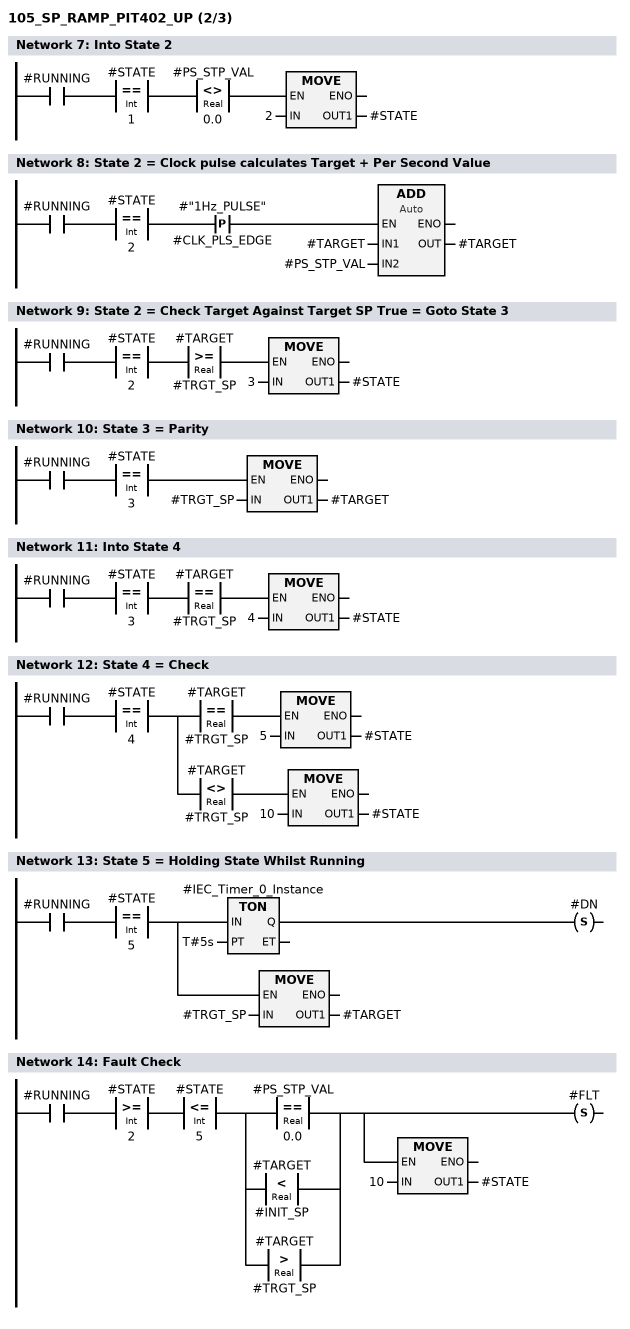
   RUNG wire#powerrail
      Contact( #RUNNING )
      { S7_Templates := "SrcType := Int" } EQ_Contact(in1 := #STATE, in2 := 1)
      { S7_Templates := "SrcType := Real" } NE_Contact(in1 := #PS_STP_VAL, in2 := 0.0)
      Move(in := 2, out1 => #STATE)
   END_RUNG
   // the same network as SCL:
   IF #RUNNING AND (#STATE = 1) AND (#PS_STP_VAL <> 0.0) THEN #STATE := 2; END_IF;
END_REGION

REGION Network 8: State 2 = Clock pulse calculates Target + Per Second Value
   RUNG wire#powerrail
      Contact( #RUNNING )
      { S7_Templates := "SrcType := Int" } EQ_Contact(in1 := #STATE, in2 := 2)
      P_Contact(operand := #"1Hz_PULSE", bit := #CLK_PLS_EDGE)
      Add(in1 := #TARGET, in2 := #PS_STP_VAL, out => #TARGET)
   END_RUNG
   // the same network as SCL:
   #_w1 := #RUNNING AND (#STATE = 2) AND #"1Hz_PULSE" AND NOT #CLK_PLS_EDGE;   // rising edge of #"1Hz_PULSE"
   #CLK_PLS_EDGE := #"1Hz_PULSE";
   IF #_w1 THEN #TARGET := #TARGET + #PS_STP_VAL; END_IF;
END_REGION

REGION Network 9: State 2 = Check Target Against Target SP True = Goto State 3
   RUNG wire#powerrail
      Contact( #RUNNING )
      { S7_Templates := "SrcType := Int" } EQ_Contact(in1 := #STATE, in2 := 2)
      { S7_Templates := "SrcType := Real" } GE_Contact(in1 := #TARGET, in2 := #TRGT_SP)
      Move(in := 3, out1 => #STATE)
   END_RUNG
   // the same network as SCL:
   IF #RUNNING AND (#STATE = 2) AND (#TARGET >= #TRGT_SP) THEN #STATE := 3; END_IF;
END_REGION

REGION Network 10: State 3 = Parity
   RUNG wire#powerrail
      Contact( #RUNNING )
      { S7_Templates := "SrcType := Int" } EQ_Contact(in1 := #STATE, in2 := 3)
      Move(in := #TRGT_SP, out1 => #TARGET)
   END_RUNG
   // the same network as SCL:
   IF #RUNNING AND (#STATE = 3) THEN #TARGET := #TRGT_SP; END_IF;
END_REGION

REGION Network 11: Into State 4
   RUNG wire#powerrail
      Contact( #RUNNING )
      { S7_Templates := "SrcType := Int" } EQ_Contact(in1 := #STATE, in2 := 3)
      { S7_Templates := "SrcType := Real" } EQ_Contact(in1 := #TARGET, in2 := #TRGT_SP)
      Move(in := 4, out1 => #STATE)
   END_RUNG
   // the same network as SCL:
   IF #RUNNING AND (#STATE = 3) AND (#TARGET = #TRGT_SP) THEN #STATE := 4; END_IF;
END_REGION

REGION Network 12: State 4 = Check
   RUNG wire#powerrail
      Contact( #RUNNING )
      { S7_Templates := "SrcType := Int" } EQ_Contact(in1 := #STATE, in2 := 4)
      wire#w1
      { S7_Templates := "SrcType := Real" } EQ_Contact(in1 := #TARGET, in2 := #TRGT_SP)
      Move(in := 5, out1 => #STATE)
   END_RUNG
   RUNG wire#w1
      { S7_Templates := "SrcType := Real" } NE_Contact(in1 := #TARGET, in2 := #TRGT_SP)
      Move(in := 10, out1 => #STATE)
   END_RUNG
   // the same network as SCL:
   #_w1 := #RUNNING AND (#STATE = 4);
   IF #_w1 AND (#TARGET = #TRGT_SP) THEN #STATE := 5; END_IF;
   IF #_w1 AND (#TARGET <> #TRGT_SP) THEN #STATE := 10; END_IF;
END_REGION

REGION Network 13: State 5 = Holding State Whilst Running
   #_w1 := #RUNNING AND (#STATE = 5);
   #IEC_Timer_0_Instance(IN := #_w1, PT := T#5s);   // TON
   IF #IEC_Timer_0_Instance.Q THEN #DN := TRUE; END_IF;
   IF #_w1 THEN #TARGET := #TRGT_SP; END_IF;
END_REGION

REGION Network 14: Fault Check
   RUNG wire#powerrail
      Contact( #RUNNING )
      { S7_Templates := "SrcType := Int" } GE_Contact(in1 := #STATE, in2 := 2)
      { S7_Templates := "SrcType := Int" } LE_Contact(in1 := #STATE, in2 := 5)
      wire#w1
      { S7_Templates := "SrcType := Real" } EQ_Contact(in1 := #PS_STP_VAL, in2 := 0.0)
      wire#w2
      S_Coil( #FLT )
   END_RUNG
   RUNG wire#w1
      { S7_Templates := "SrcType := Real" } LT_Contact(in1 := #TARGET, in2 := #INIT_SP)
   END_RUNG wire#w2
   RUNG wire#w1
      { S7_Templates := "SrcType := Real" } GT_Contact(in1 := #TARGET, in2 := #TRGT_SP)
   END_RUNG wire#w2
   RUNG wire#w2
      Move(in := 10, out1 => #STATE)
   END_RUNG
   // the same network as SCL:
   IF #RUNNING AND (#STATE >= 2) AND (#STATE <= 5) AND ((#PS_STP_VAL = 0.0) OR (#TARGET < #INIT_SP) OR (#TARGET > #TRGT_SP)) THEN
       #FLT := TRUE;
       #STATE := 10;
   END_IF;
END_REGION

REGION Network 15: State 10 = Fault
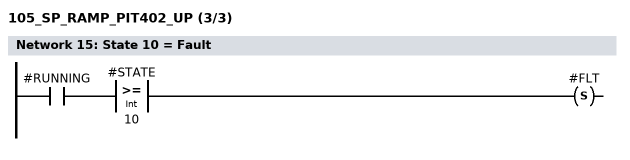
   RUNG wire#powerrail
      Contact( #RUNNING )
      { S7_Templates := "SrcType := Int" } GE_Contact(in1 := #STATE, in2 := 10)
      S_Coil( #FLT )
   END_RUNG
   // the same network as SCL:
   IF #RUNNING AND (#STATE >= 10) THEN #FLT := TRUE; END_IF;
END_REGION
END_FUNCTION_BLOCK

FUNCTION_BLOCK "107_SP_RAMP_PIT402_DN"   // FB107, LAD
TITLE = Setpoint Ramp Down For PIT402
{ S7_Optimized_Access := 'TRUE' }
AUTHOR : JRS
VERSION : 0.1
// Determines the live setpoint value for PIT402 based on target and ramp time
   VAR_INPUT
      RUN : Bool;   // Demand
      INIT_SP : Real;   // Initial setpoint
      TRGT_SP : Real;   // Target setpoint
      RMP_SECS : Int := 30;   // To target ramp time in seconds
      "1Hz_PULSE" : Bool;   // 1 Hz clock pulse
      RST : Bool;   // Reset flag
   END_VAR
   VAR_OUTPUT
      DN : Bool;   // Done
      FLT : Bool;   // Fault
   END_VAR
   VAR_IN_OUT
      RUNNING : Bool;   // Block is running
      TARGET : Real;   // Target
   END_VAR
   VAR
      STATE : Int;   // State value
      INTO_RUN_EDGE : Bool;   // Edge bit
      OUT_OF_RUN_EDGE : Bool;   // Edge bit
      RST_FLG : Bool;   // Reset flag
      PS_STP_VAL : Real;   // Per second step value
      CLK_PLS_EDGE : Bool;   // Clock pulse edge
   END_VAR
   VAR_TEMP   // added for the SCL form of the ladder/FBD networks
      _w1 : Bool;
   END_VAR
BEGIN

REGION Network 1: Running
   // For running status detection
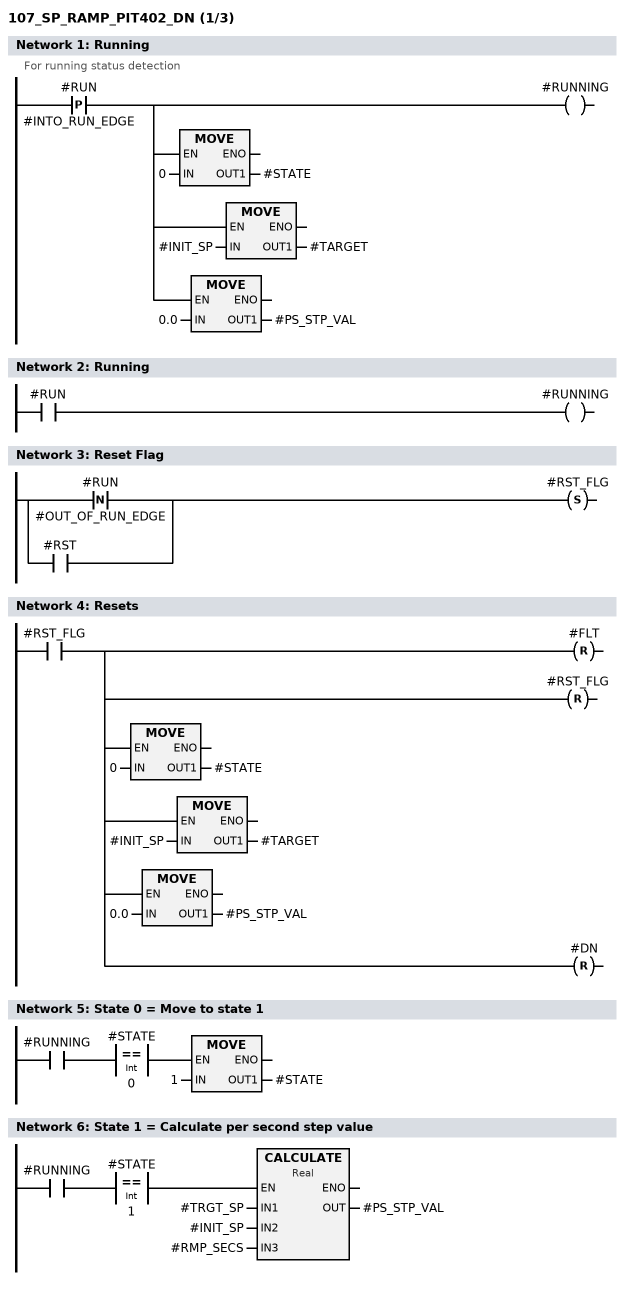
   RUNG wire#powerrail
      P_Contact(operand := #RUN, bit := #INTO_RUN_EDGE)
      wire#w1
      Coil( #RUNNING )
   END_RUNG
   RUNG wire#w1
      Move(in := 0, out1 => #STATE)
   END_RUNG
   RUNG wire#w1
      Move(in := #INIT_SP, out1 => #TARGET)
   END_RUNG
   RUNG wire#w1
      Move(in := 0.0, out1 => #PS_STP_VAL)
   END_RUNG
   // the same network as SCL:
   #_w1 := #RUN AND NOT #INTO_RUN_EDGE;   // rising edge of #RUN
   #INTO_RUN_EDGE := #RUN;
   #RUNNING := #_w1;
   IF #_w1 THEN
       #STATE := 0;
       #TARGET := #INIT_SP;
       #PS_STP_VAL := 0.0;
   END_IF;
END_REGION

REGION Network 2: Running
   RUNG wire#powerrail
      Contact( #RUN )
      Coil( #RUNNING )
   END_RUNG
   // the same network as SCL:
   #RUNNING := #RUN;
END_REGION

REGION Network 3: Reset Flag
   RUNG wire#powerrail
      N_Contact(operand := #RUN, bit := #OUT_OF_RUN_EDGE)
      wire#w1
      S_Coil( #RST_FLG )
   END_RUNG
   RUNG wire#powerrail
      Contact( #RST )
   END_RUNG wire#w1
   // the same network as SCL:
   #_w1 := NOT #RUN AND #OUT_OF_RUN_EDGE;   // falling edge of #RUN
   #OUT_OF_RUN_EDGE := #RUN;
   IF #_w1 OR #RST THEN #RST_FLG := TRUE; END_IF;
END_REGION

REGION Network 4: Resets
   RUNG wire#powerrail
      Contact( #RST_FLG )
      wire#w1
      R_Coil( #FLT )
   END_RUNG
   RUNG wire#w1
      R_Coil( #RST_FLG )
   END_RUNG
   RUNG wire#w1
      Move(in := 0, out1 => #STATE)
   END_RUNG
   RUNG wire#w1
      Move(in := #INIT_SP, out1 => #TARGET)
   END_RUNG
   RUNG wire#w1
      Move(in := 0.0, out1 => #PS_STP_VAL)
   END_RUNG
   RUNG wire#w1
      R_Coil( #DN )
   END_RUNG
   // the same network as SCL:
   IF #RST_FLG THEN #FLT := FALSE; END_IF;
   #_w1 := #RST_FLG;
   IF #_w1 THEN
       #RST_FLG := FALSE;
       #STATE := 0;
       #TARGET := #INIT_SP;
       #PS_STP_VAL := 0.0;
       #DN := FALSE;
   END_IF;
END_REGION

REGION Network 5: State 0 = Move to state 1
   RUNG wire#powerrail
      Contact( #RUNNING )
      { S7_Templates := "SrcType := Int" } EQ_Contact(in1 := #STATE, in2 := 0)
      Move(in := 1, out1 => #STATE)
   END_RUNG
   // the same network as SCL:
   IF #RUNNING AND (#STATE = 0) THEN #STATE := 1; END_IF;
END_REGION

REGION Network 6: State 1 = Calculate per second step value
   RUNG wire#powerrail
      Contact( #RUNNING )
      { S7_Templates := "SrcType := Int" } EQ_Contact(in1 := #STATE, in2 := 1)
      { S7_Templates := "SrcType := Real"; S7_Expression := "(IN2-IN1)/IN3" } Calculate(in1 := #TRGT_SP, in2 := #INIT_SP, in3 := #RMP_SECS, out => #PS_STP_VAL)
   END_RUNG
   // the same network as SCL:
   IF #RUNNING AND (#STATE = 1) THEN #PS_STP_VAL := (#INIT_SP-#TRGT_SP)/#RMP_SECS; END_IF;
END_REGION

REGION Network 7: Into State 2
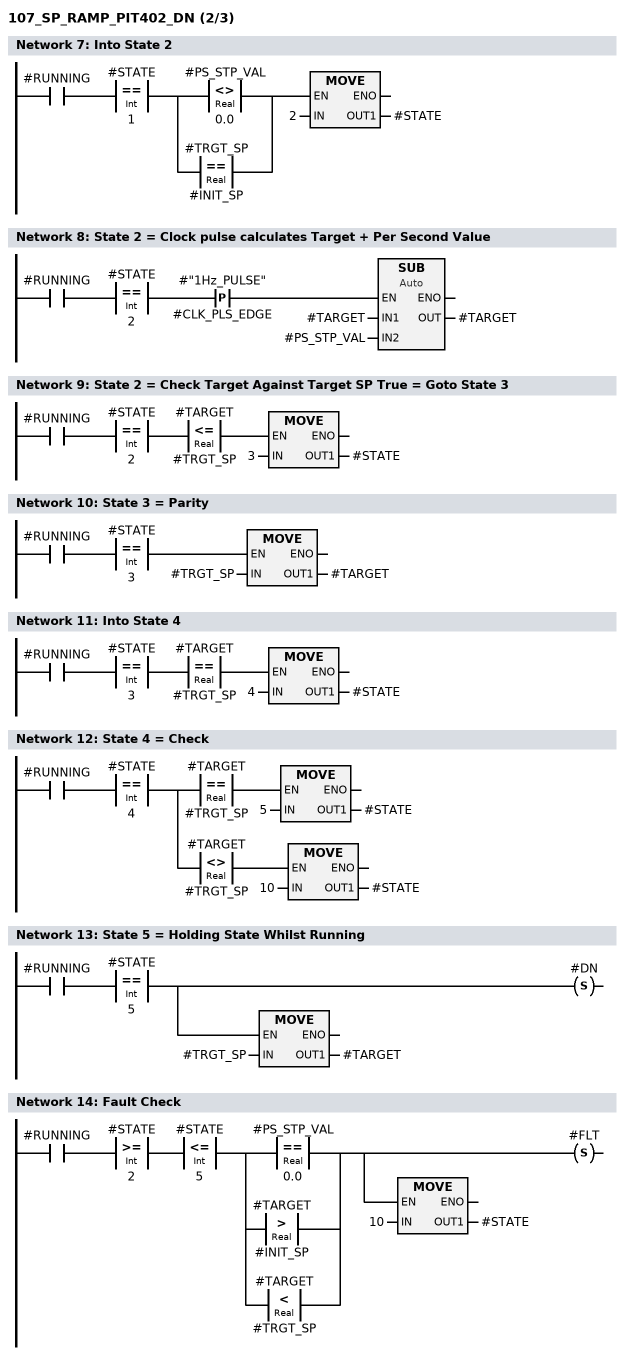
   RUNG wire#powerrail
      Contact( #RUNNING )
      { S7_Templates := "SrcType := Int" } EQ_Contact(in1 := #STATE, in2 := 1)
      wire#w1
      { S7_Templates := "SrcType := Real" } NE_Contact(in1 := #PS_STP_VAL, in2 := 0.0)
      wire#w2
      Move(in := 2, out1 => #STATE)
   END_RUNG
   RUNG wire#w1
      { S7_Templates := "SrcType := Real" } EQ_Contact(in1 := #TRGT_SP, in2 := #INIT_SP)
   END_RUNG wire#w2
   // the same network as SCL:
   IF #RUNNING AND (#STATE = 1) AND ((#PS_STP_VAL <> 0.0) OR (#TRGT_SP = #INIT_SP)) THEN #STATE := 2; END_IF;
END_REGION

REGION Network 8: State 2 = Clock pulse calculates Target + Per Second Value
   RUNG wire#powerrail
      Contact( #RUNNING )
      { S7_Templates := "SrcType := Int" } EQ_Contact(in1 := #STATE, in2 := 2)
      P_Contact(operand := #"1Hz_PULSE", bit := #CLK_PLS_EDGE)
      Sub(in1 := #TARGET, in2 := #PS_STP_VAL, out => #TARGET)
   END_RUNG
   // the same network as SCL:
   #_w1 := #RUNNING AND (#STATE = 2) AND #"1Hz_PULSE" AND NOT #CLK_PLS_EDGE;   // rising edge of #"1Hz_PULSE"
   #CLK_PLS_EDGE := #"1Hz_PULSE";
   IF #_w1 THEN #TARGET := #TARGET - #PS_STP_VAL; END_IF;
END_REGION

REGION Network 9: State 2 = Check Target Against Target SP True = Goto State 3
   RUNG wire#powerrail
      Contact( #RUNNING )
      { S7_Templates := "SrcType := Int" } EQ_Contact(in1 := #STATE, in2 := 2)
      { S7_Templates := "SrcType := Real" } LE_Contact(in1 := #TARGET, in2 := #TRGT_SP)
      Move(in := 3, out1 => #STATE)
   END_RUNG
   // the same network as SCL:
   IF #RUNNING AND (#STATE = 2) AND (#TARGET <= #TRGT_SP) THEN #STATE := 3; END_IF;
END_REGION

REGION Network 10: State 3 = Parity
   RUNG wire#powerrail
      Contact( #RUNNING )
      { S7_Templates := "SrcType := Int" } EQ_Contact(in1 := #STATE, in2 := 3)
      Move(in := #TRGT_SP, out1 => #TARGET)
   END_RUNG
   // the same network as SCL:
   IF #RUNNING AND (#STATE = 3) THEN #TARGET := #TRGT_SP; END_IF;
END_REGION

REGION Network 11: Into State 4
   RUNG wire#powerrail
      Contact( #RUNNING )
      { S7_Templates := "SrcType := Int" } EQ_Contact(in1 := #STATE, in2 := 3)
      { S7_Templates := "SrcType := Real" } EQ_Contact(in1 := #TARGET, in2 := #TRGT_SP)
      Move(in := 4, out1 => #STATE)
   END_RUNG
   // the same network as SCL:
   IF #RUNNING AND (#STATE = 3) AND (#TARGET = #TRGT_SP) THEN #STATE := 4; END_IF;
END_REGION

REGION Network 12: State 4 = Check
   RUNG wire#powerrail
      Contact( #RUNNING )
      { S7_Templates := "SrcType := Int" } EQ_Contact(in1 := #STATE, in2 := 4)
      wire#w1
      { S7_Templates := "SrcType := Real" } EQ_Contact(in1 := #TARGET, in2 := #TRGT_SP)
      Move(in := 5, out1 => #STATE)
   END_RUNG
   RUNG wire#w1
      { S7_Templates := "SrcType := Real" } NE_Contact(in1 := #TARGET, in2 := #TRGT_SP)
      Move(in := 10, out1 => #STATE)
   END_RUNG
   // the same network as SCL:
   #_w1 := #RUNNING AND (#STATE = 4);
   IF #_w1 AND (#TARGET = #TRGT_SP) THEN #STATE := 5; END_IF;
   IF #_w1 AND (#TARGET <> #TRGT_SP) THEN #STATE := 10; END_IF;
END_REGION

REGION Network 13: State 5 = Holding State Whilst Running
   RUNG wire#powerrail
      Contact( #RUNNING )
      { S7_Templates := "SrcType := Int" } EQ_Contact(in1 := #STATE, in2 := 5)
      wire#w1
      S_Coil( #DN )
   END_RUNG
   RUNG wire#w1
      Move(in := #TRGT_SP, out1 => #TARGET)
   END_RUNG
   // the same network as SCL:
   IF #RUNNING AND (#STATE = 5) THEN
       #DN := TRUE;
       #TARGET := #TRGT_SP;
   END_IF;
END_REGION

REGION Network 14: Fault Check
   RUNG wire#powerrail
      Contact( #RUNNING )
      { S7_Templates := "SrcType := Int" } GE_Contact(in1 := #STATE, in2 := 2)
      { S7_Templates := "SrcType := Int" } LE_Contact(in1 := #STATE, in2 := 5)
      wire#w1
      { S7_Templates := "SrcType := Real" } EQ_Contact(in1 := #PS_STP_VAL, in2 := 0.0)
      wire#w2
      S_Coil( #FLT )
   END_RUNG
   RUNG wire#w1
      { S7_Templates := "SrcType := Real" } GT_Contact(in1 := #TARGET, in2 := #INIT_SP)
   END_RUNG wire#w2
   RUNG wire#w1
      { S7_Templates := "SrcType := Real" } LT_Contact(in1 := #TARGET, in2 := #TRGT_SP)
   END_RUNG wire#w2
   RUNG wire#w2
      Move(in := 10, out1 => #STATE)
   END_RUNG
   // the same network as SCL:
   IF #RUNNING AND (#STATE >= 2) AND (#STATE <= 5) AND ((#PS_STP_VAL = 0.0) OR (#TARGET > #INIT_SP) OR (#TARGET < #TRGT_SP)) THEN
       #FLT := TRUE;
       #STATE := 10;
   END_IF;
END_REGION

REGION Network 15: State 10 = Fault
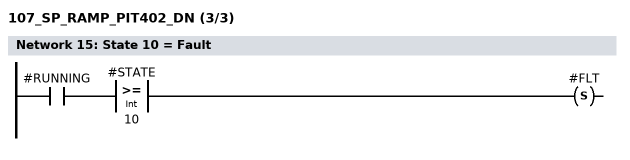
   RUNG wire#powerrail
      Contact( #RUNNING )
      { S7_Templates := "SrcType := Int" } GE_Contact(in1 := #STATE, in2 := 10)
      S_Coil( #FLT )
   END_RUNG
   // the same network as SCL:
   IF #RUNNING AND (#STATE >= 10) THEN #FLT := TRUE; END_IF;
END_REGION
END_FUNCTION_BLOCK

FUNCTION "100_SC" : Void   // FC100, LAD
TITLE = State Complete
{ S7_Optimized_Access := 'TRUE' }
AUTHOR : JRS
VERSION : 0.1
// For the determination of each step state being complete
   VAR_TEMP   // added for the SCL form of the ladder/FBD networks
      _w1 : Bool;
   END_VAR
BEGIN

REGION Network 1: Step 001 = Confirm Auto Conditions Ok
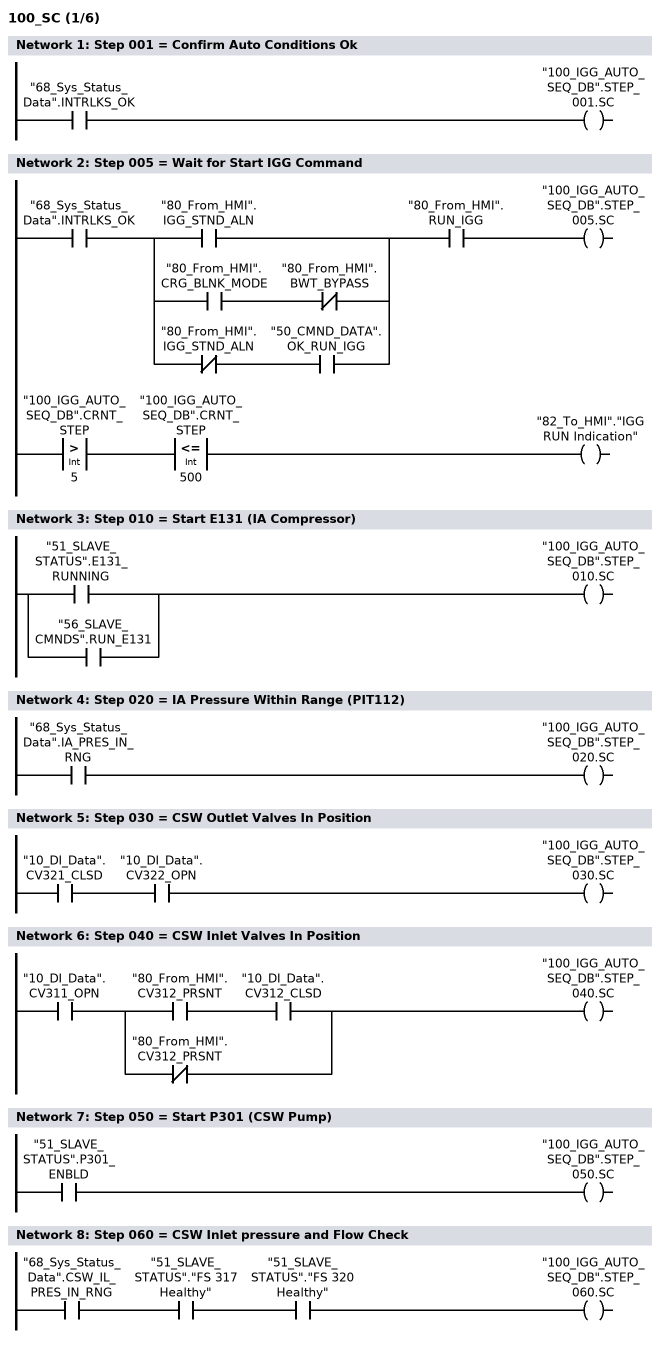
   RUNG wire#powerrail
      Contact( "68_Sys_Status_Data".INTRLKS_OK )
      Coil( "100_IGG_AUTO_SEQ_DB".STEP_001.SC )
   END_RUNG
   // the same network as SCL:
   "100_IGG_AUTO_SEQ_DB".STEP_001.SC := "68_Sys_Status_Data".INTRLKS_OK;
END_REGION

REGION Network 2: Step 005 = Wait for Start IGG Command
   RUNG wire#powerrail
      Contact( "68_Sys_Status_Data".INTRLKS_OK )
      wire#w1
      Contact( "80_From_HMI".IGG_STND_ALN )
      wire#w2
      Contact( "80_From_HMI".RUN_IGG )
      Coil( "100_IGG_AUTO_SEQ_DB".STEP_005.SC )
   END_RUNG
   RUNG wire#w1
      Contact( "80_From_HMI".CRG_BLNK_MODE )
      I_Contact( "80_From_HMI".BWT_BYPASS )
   END_RUNG wire#w2
   RUNG wire#w1
      I_Contact( "80_From_HMI".IGG_STND_ALN )
      Contact( "50_CMND_DATA".OK_RUN_IGG )
   END_RUNG wire#w2
   RUNG wire#powerrail
      { S7_Templates := "SrcType := Int" } GT_Contact(in1 := "100_IGG_AUTO_SEQ_DB".CRNT_STEP, in2 := 5)
      { S7_Templates := "SrcType := Int" } LE_Contact(in1 := "100_IGG_AUTO_SEQ_DB".CRNT_STEP, in2 := 500)
      Coil( "82_To_HMI"."IGG RUN Indication" )
   END_RUNG
   // the same network as SCL:
   "100_IGG_AUTO_SEQ_DB".STEP_005.SC := "68_Sys_Status_Data".INTRLKS_OK AND ("80_From_HMI".IGG_STND_ALN OR ("80_From_HMI".CRG_BLNK_MODE AND NOT "80_From_HMI".BWT_BYPASS) OR (NOT "80_From_HMI".IGG_STND_ALN AND "50_CMND_DATA".OK_RUN_IGG)) AND "80_From_HMI".RUN_IGG;
   "82_To_HMI"."IGG RUN Indication" := ("100_IGG_AUTO_SEQ_DB".CRNT_STEP > 5) AND ("100_IGG_AUTO_SEQ_DB".CRNT_STEP <= 500);
END_REGION

REGION Network 3: Step 010 = Start E131 (IA Compressor)
   RUNG wire#powerrail
      Contact( "51_SLAVE_STATUS".E131_RUNNING )
      wire#w1
      Coil( "100_IGG_AUTO_SEQ_DB".STEP_010.SC )
   END_RUNG
   RUNG wire#powerrail
      Contact( "56_SLAVE_CMNDS".RUN_E131 )
   END_RUNG wire#w1
   // the same network as SCL:
   "100_IGG_AUTO_SEQ_DB".STEP_010.SC := "51_SLAVE_STATUS".E131_RUNNING OR "56_SLAVE_CMNDS".RUN_E131;
END_REGION

REGION Network 4: Step 020 = IA Pressure Within Range (PIT112)
   RUNG wire#powerrail
      Contact( "68_Sys_Status_Data".IA_PRES_IN_RNG )
      Coil( "100_IGG_AUTO_SEQ_DB".STEP_020.SC )
   END_RUNG
   // the same network as SCL:
   "100_IGG_AUTO_SEQ_DB".STEP_020.SC := "68_Sys_Status_Data".IA_PRES_IN_RNG;
END_REGION

REGION Network 5: Step 030 = CSW Outlet Valves In Position
   RUNG wire#powerrail
      Contact( "10_DI_Data".CV321_CLSD )
      Contact( "10_DI_Data".CV322_OPN )
      Coil( "100_IGG_AUTO_SEQ_DB".STEP_030.SC )
   END_RUNG
   // the same network as SCL:
   "100_IGG_AUTO_SEQ_DB".STEP_030.SC := "10_DI_Data".CV321_CLSD AND "10_DI_Data".CV322_OPN;
END_REGION

REGION Network 6: Step 040 = CSW Inlet Valves In Position
   RUNG wire#powerrail
      Contact( "10_DI_Data".CV311_OPN )
      wire#w1
      Contact( "80_From_HMI".CV312_PRSNT )
      Contact( "10_DI_Data".CV312_CLSD )
      wire#w2
      Coil( "100_IGG_AUTO_SEQ_DB".STEP_040.SC )
   END_RUNG
   RUNG wire#w1
      I_Contact( "80_From_HMI".CV312_PRSNT )
   END_RUNG wire#w2
   // the same network as SCL:
   "100_IGG_AUTO_SEQ_DB".STEP_040.SC := "10_DI_Data".CV311_OPN AND (("80_From_HMI".CV312_PRSNT AND "10_DI_Data".CV312_CLSD) OR NOT "80_From_HMI".CV312_PRSNT);
END_REGION

REGION Network 7: Step 050 = Start P301 (CSW Pump)
   RUNG wire#powerrail
      Contact( "51_SLAVE_STATUS".P301_ENBLD )
      Coil( "100_IGG_AUTO_SEQ_DB".STEP_050.SC )
   END_RUNG
   // the same network as SCL:
   "100_IGG_AUTO_SEQ_DB".STEP_050.SC := "51_SLAVE_STATUS".P301_ENBLD;
END_REGION

REGION Network 8: Step 060 = CSW Inlet pressure and Flow Check
   RUNG wire#powerrail
      Contact( "68_Sys_Status_Data".CSW_IL_PRES_IN_RNG )
      Contact( "51_SLAVE_STATUS"."FS 317 Healthy" )
      Contact( "51_SLAVE_STATUS"."FS 320 Healthy" )
      Coil( "100_IGG_AUTO_SEQ_DB".STEP_060.SC )
   END_RUNG
   // the same network as SCL:
   "100_IGG_AUTO_SEQ_DB".STEP_060.SC := "68_Sys_Status_Data".CSW_IL_PRES_IN_RNG AND "51_SLAVE_STATUS"."FS 317 Healthy" AND "51_SLAVE_STATUS"."FS 320 Healthy";
END_REGION

REGION Network 9: Step 070 = Check CV203 Position Closed (N.C.)
   // This valve is on the BC PLC with no tell-back
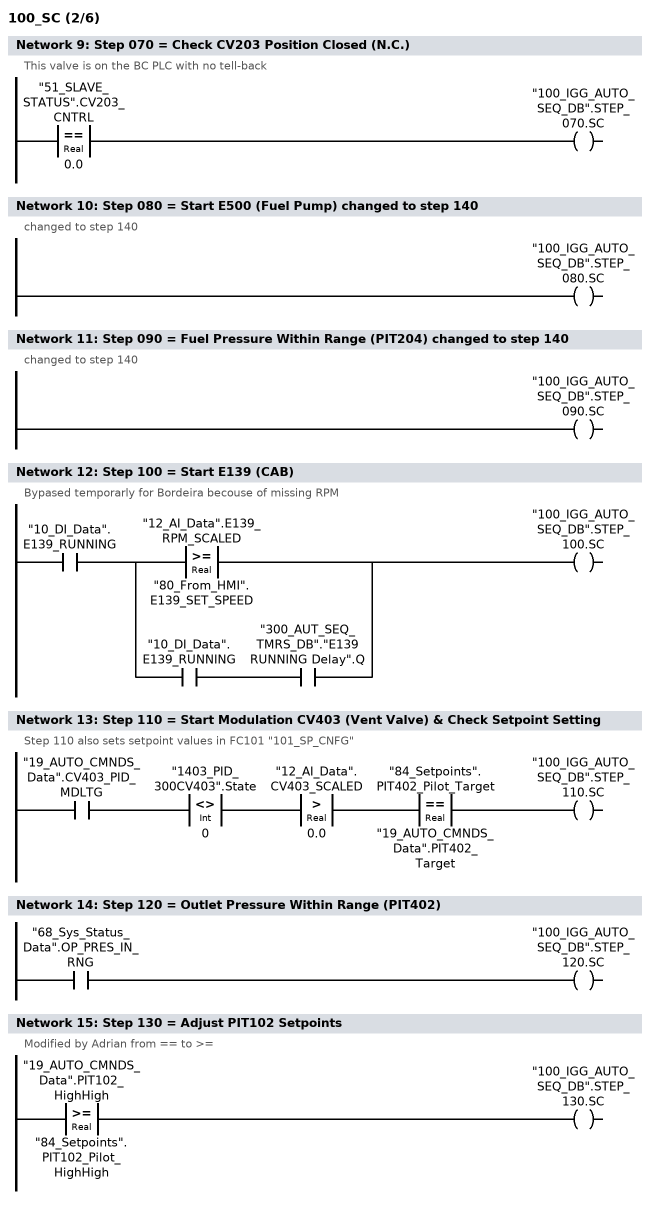
   RUNG wire#powerrail
      { S7_Templates := "SrcType := Real" } EQ_Contact(in1 := "51_SLAVE_STATUS".CV203_CNTRL, in2 := 0.0)
      Coil( "100_IGG_AUTO_SEQ_DB".STEP_070.SC )
   END_RUNG
   // the same network as SCL:
   "100_IGG_AUTO_SEQ_DB".STEP_070.SC := "51_SLAVE_STATUS".CV203_CNTRL = 0.0;
END_REGION

REGION Network 10: Step 080 = Start E500 (Fuel Pump) changed to step 140
   // changed to step 140
   RUNG wire#powerrail
      Coil( "100_IGG_AUTO_SEQ_DB".STEP_080.SC )
   END_RUNG
   // the same network as SCL:
   "100_IGG_AUTO_SEQ_DB".STEP_080.SC := TRUE;
END_REGION

REGION Network 11: Step 090 = Fuel Pressure Within Range (PIT204) changed to step 140
   // changed to step 140
   RUNG wire#powerrail
      Coil( "100_IGG_AUTO_SEQ_DB".STEP_090.SC )
   END_RUNG
   // the same network as SCL:
   "100_IGG_AUTO_SEQ_DB".STEP_090.SC := TRUE;
END_REGION

REGION Network 12: Step 100 = Start E139 (CAB)
   // Bypased temporarly for Bordeira becouse of missing RPM
   RUNG wire#powerrail
      Contact( "10_DI_Data".E139_RUNNING )
      wire#w1
      { S7_Templates := "SrcType := Real" } GE_Contact(in1 := "12_AI_Data".E139_RPM_SCALED, in2 := "80_From_HMI".E139_SET_SPEED)
      wire#w2
      Coil( "100_IGG_AUTO_SEQ_DB".STEP_100.SC )
   END_RUNG
   RUNG wire#w1
      Contact( "10_DI_Data".E139_RUNNING )
      Contact( "300_AUT_SEQ_TMRS_DB"."E139 RUNNING Delay".Q )
   END_RUNG wire#w2
   // the same network as SCL:
   "100_IGG_AUTO_SEQ_DB".STEP_100.SC := "10_DI_Data".E139_RUNNING AND (("12_AI_Data".E139_RPM_SCALED >= "80_From_HMI".E139_SET_SPEED) OR ("10_DI_Data".E139_RUNNING AND "300_AUT_SEQ_TMRS_DB"."E139 RUNNING Delay".Q));
END_REGION

REGION Network 13: Step 110 = Start Modulation CV403 (Vent Valve) & Check Setpoint Setting
   // Step 110 also sets setpoint values in FC101 "101_SP_CNFG"
   RUNG wire#powerrail
      Contact( "19_AUTO_CMNDS_Data".CV403_PID_MDLTG )
      { S7_Templates := "SrcType := Int" } NE_Contact(in1 := "1403_PID_300CV403".State, in2 := 0)
      { S7_Templates := "SrcType := Real" } GT_Contact(in1 := "12_AI_Data".CV403_SCALED, in2 := 0.0)
      { S7_Templates := "SrcType := Real" } EQ_Contact(in1 := "84_Setpoints".PIT402_Pilot_Target, in2 := "19_AUTO_CMNDS_Data".PIT402_Target)
      Coil( "100_IGG_AUTO_SEQ_DB".STEP_110.SC )
   END_RUNG
   // the same network as SCL:
   "100_IGG_AUTO_SEQ_DB".STEP_110.SC := "19_AUTO_CMNDS_Data".CV403_PID_MDLTG AND ("1403_PID_300CV403".State <> 0) AND ("12_AI_Data".CV403_SCALED > 0.0) AND ("84_Setpoints".PIT402_Pilot_Target = "19_AUTO_CMNDS_Data".PIT402_Target);
END_REGION

REGION Network 14: Step 120 = Outlet Pressure Within Range (PIT402)
   RUNG wire#powerrail
      Contact( "68_Sys_Status_Data".OP_PRES_IN_RNG )
      Coil( "100_IGG_AUTO_SEQ_DB".STEP_120.SC )
   END_RUNG
   // the same network as SCL:
   "100_IGG_AUTO_SEQ_DB".STEP_120.SC := "68_Sys_Status_Data".OP_PRES_IN_RNG;
END_REGION

REGION Network 15: Step 130 = Adjust PIT102 Setpoints
   // Modified by Adrian from == to >=
   RUNG wire#powerrail
      { S7_Templates := "SrcType := Real" } GE_Contact(in1 := "19_AUTO_CMNDS_Data".PIT102_HighHigh, in2 := "84_Setpoints".PIT102_Pilot_HighHigh)
      Coil( "100_IGG_AUTO_SEQ_DB".STEP_130.SC )
   END_RUNG
   // the same network as SCL:
   "100_IGG_AUTO_SEQ_DB".STEP_130.SC := "19_AUTO_CMNDS_Data".PIT102_HighHigh >= "84_Setpoints".PIT102_Pilot_HighHigh;
END_REGION

REGION Network 16: Step 140 = Pre BC Start Sequence Delay
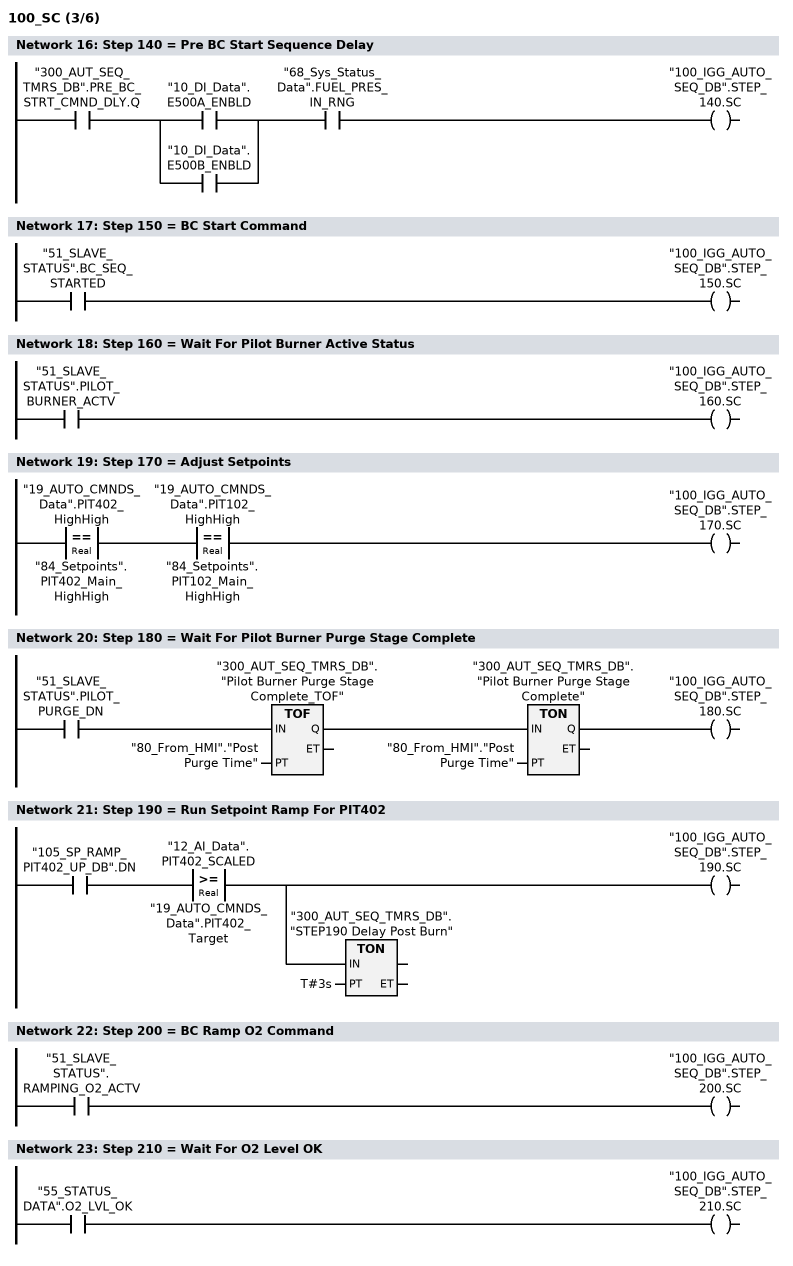
   RUNG wire#powerrail
      Contact( "300_AUT_SEQ_TMRS_DB".PRE_BC_STRT_CMND_DLY.Q )
      wire#w1
      Contact( "10_DI_Data".E500A_ENBLD )
      wire#w2
      Contact( "68_Sys_Status_Data".FUEL_PRES_IN_RNG )
      Coil( "100_IGG_AUTO_SEQ_DB".STEP_140.SC )
   END_RUNG
   RUNG wire#w1
      Contact( "10_DI_Data".E500B_ENBLD )
   END_RUNG wire#w2
   // the same network as SCL:
   "100_IGG_AUTO_SEQ_DB".STEP_140.SC := "300_AUT_SEQ_TMRS_DB".PRE_BC_STRT_CMND_DLY.Q AND ("10_DI_Data".E500A_ENBLD OR "10_DI_Data".E500B_ENBLD) AND "68_Sys_Status_Data".FUEL_PRES_IN_RNG;
END_REGION

REGION Network 17: Step 150 = BC Start Command
   RUNG wire#powerrail
      Contact( "51_SLAVE_STATUS".BC_SEQ_STARTED )
      Coil( "100_IGG_AUTO_SEQ_DB".STEP_150.SC )
   END_RUNG
   // the same network as SCL:
   "100_IGG_AUTO_SEQ_DB".STEP_150.SC := "51_SLAVE_STATUS".BC_SEQ_STARTED;
END_REGION

REGION Network 18: Step 160 = Wait For Pilot Burner Active Status
   RUNG wire#powerrail
      Contact( "51_SLAVE_STATUS".PILOT_BURNER_ACTV )
      Coil( "100_IGG_AUTO_SEQ_DB".STEP_160.SC )
   END_RUNG
   // the same network as SCL:
   "100_IGG_AUTO_SEQ_DB".STEP_160.SC := "51_SLAVE_STATUS".PILOT_BURNER_ACTV;
END_REGION

REGION Network 19: Step 170 = Adjust Setpoints
   RUNG wire#powerrail
      { S7_Templates := "SrcType := Real" } EQ_Contact(in1 := "19_AUTO_CMNDS_Data".PIT402_HighHigh, in2 := "84_Setpoints".PIT402_Main_HighHigh)
      { S7_Templates := "SrcType := Real" } EQ_Contact(in1 := "19_AUTO_CMNDS_Data".PIT102_HighHigh, in2 := "84_Setpoints".PIT102_Main_HighHigh)
      Coil( "100_IGG_AUTO_SEQ_DB".STEP_170.SC )
   END_RUNG
   // the same network as SCL:
   "100_IGG_AUTO_SEQ_DB".STEP_170.SC := ("19_AUTO_CMNDS_Data".PIT402_HighHigh = "84_Setpoints".PIT402_Main_HighHigh) AND ("19_AUTO_CMNDS_Data".PIT102_HighHigh = "84_Setpoints".PIT102_Main_HighHigh);
END_REGION

REGION Network 20: Step 180 = Wait For Pilot Burner Purge Stage Complete
   "300_AUT_SEQ_TMRS_DB"."Pilot Burner Purge Stage Complete_TOF".TOF(IN := "51_SLAVE_STATUS".PILOT_PURGE_DN,
                           PT := "80_From_HMI"."Post Purge Time");
   "300_AUT_SEQ_TMRS_DB"."Pilot Burner Purge Stage Complete".TON(IN := "300_AUT_SEQ_TMRS_DB"."Pilot Burner Purge Stage Complete_TOF".Q,
                           PT := "80_From_HMI"."Post Purge Time");
   "100_IGG_AUTO_SEQ_DB".STEP_180.SC := "300_AUT_SEQ_TMRS_DB"."Pilot Burner Purge Stage Complete".Q;
END_REGION

REGION Network 21: Step 190 = Run Setpoint Ramp For PIT402
   "100_IGG_AUTO_SEQ_DB".STEP_190.SC := "105_SP_RAMP_PIT402_UP_DB".DN AND ("12_AI_Data".PIT402_SCALED >= "19_AUTO_CMNDS_Data".PIT402_Target);
   "300_AUT_SEQ_TMRS_DB"."STEP190 Delay Post Burn".TON(IN := "100_IGG_AUTO_SEQ_DB".STEP_190.SC, PT := T#3s);
END_REGION

REGION Network 22: Step 200 = BC Ramp O2 Command
   RUNG wire#powerrail
      Contact( "51_SLAVE_STATUS".RAMPING_O2_ACTV )
      Coil( "100_IGG_AUTO_SEQ_DB".STEP_200.SC )
   END_RUNG
   // the same network as SCL:
   "100_IGG_AUTO_SEQ_DB".STEP_200.SC := "51_SLAVE_STATUS".RAMPING_O2_ACTV;
END_REGION

REGION Network 23: Step 210 = Wait For O2 Level OK
   RUNG wire#powerrail
      Contact( "55_STATUS_DATA".O2_LVL_OK )
      Coil( "100_IGG_AUTO_SEQ_DB".STEP_210.SC )
   END_RUNG
   // the same network as SCL:
   "100_IGG_AUTO_SEQ_DB".STEP_210.SC := "55_STATUS_DATA".O2_LVL_OK;
END_REGION

REGION Network 24: Step 220 = Wait For Stop Command